HMI tags "New_Added"
   "AbufferCopyCut" : Bool, internal
   "AbufferFile" : WString[255], internal
   "AbufferFolder" : WString[255], internal
   "AbufferIsFolder" : Bool, internal
   "AFEsearchFolder" : WString[80], internal
   "AFEsearchString" : WString[80], internal
   "AFEStatus" : WString[150], internal
   "AFile_1" : WString[255], internal
   "AFile_10" : WString[255], internal
   "AFile_2" : WString[255], internal
   "AFile_3" : WString[255], internal
   "AFile_4" : WString[255], internal
   "AFile_5" : WString[255], internal
   "AFile_6" : WString[255], internal
   "AFile_7" : WString[255], internal
   "AFile_8" : WString[255], internal
   "AFile_9" : WString[255], internal
   "AfileChosen" : Int, internal
   "AFolder" : WString[255], internal
   "AhtmlPath" : WString[80], internal
   "Aindex" : Int, internal
   "AisFolder_1" : WString[10], internal
   "AisFolder_10" : WString[10], internal
   "AisFolder_2" : WString[10], internal
   "AisFolder_3" : WString[10], internal
   "AisFolder_4" : WString[10], internal
   "AisFolder_5" : WString[10], internal
   "AisFolder_6" : WString[10], internal
   "AisFolder_7" : WString[10], internal
   "AisFolder_8" : WString[10], internal
   "AisFolder_9" : WString[10], internal
   "ANewFolder" : WString[255], internal
   "ANewName" : WString[255], internal
   "ANextPossible" : Bool, internal
   "ApdfPath" : WString[80], internal
   "ASearch" : Bool, internal
   "AstateBackground" : Bool, internal
   "copyusb" : Bool, internal

HMI tags "NEW"
   "PV_1" : DInt AT %DB12.DBD32, 1 s
   "PV_2" : DInt AT %DB13.DBD28, 1 s
   "PV_3" : Int AT %DB12.DBW6, 1 s
   "SV_1" : DInt AT %DB16.DBD26, 1 s
   "SV_2" : Int AT %DB14.DBW20, 1 s
   "SV_3" : Int AT %DB12.DBW4, 1 s
   "Selection" : Bool AT %M30.0, 1 s
   "F2" : Bool AT %M30.1, 1 s
   "F3" : Bool AT %M33.3, 1 s
   "F4" : Bool AT %M33.4, 1 s
   "F5" : Bool AT %M30.3, 1 s
   "ON_OFF" : Bool AT %M30.1, 1 s
   "Indicator" : Bool AT %Q124.2, 1 s
   "F6" : Bool AT %M30.4, 1 s

discrete alarms
   1: 'All logs have been closed successfully.', class Sampling, trigger "Sampling_Alarm" bit 0
      on Coming: function_a9b64e44("Sampling_Alarm", 0)
   2: 'Log initialization ended. All logs OK.', class Sampling, trigger "Sampling_Alarm" bit 1
      on Coming: function_a9b64e44("Sampling_Alarm", 1)
   3: 'The log was successfully exported / The log was successfully exported to SD Card', class Sampling, trigger "Sampling_Alarm" bit 2
      on Coming: function_a9b64e44("Sampling_Alarm", 2)

text list "FLow_RPM": 0 'RPM'; 1 'FLOW RATE'

text list "ON_OFF": 0 'OFF'; 1 'ON'

graphic list "Nav_Recipe": 0 'labu1'; 1 'labu2'

graphic list "Check_Uncheck": 0 'images (7)'; 1 '_green_check.svg'

graphic list "pump": 2 'motor2'; 1 'motor'; 3 'motor'; 4 'motor2'; 5 'motor'; 6 'motor2'

graphic list "MH": 0 'graph'; 1 'graph - Copy'

graphic list "Home": 0 'images_3'; 1 'images - Copy'

graphic list "Scope": 0..12 'scope_1'; 13 'scope - Copy'; 14 'scope_1'

graphic list "oscilloscope": 0..8 'osiloskope'; 9 'osiloskope - Copy'; 10..14 'osiloskope'

graphic list "SelectorMenu": 0..10 's2_1'; 11 's2 - Copy'; 12..14 's2_1'

graphic list "Color": 0 'color1'; 1 'color1'; 2 'color3'; 4 'color5'; 8 'color6'; 16 'color7'

graphic list "SettingSys1": 0..6 'settingsys_1'; 7..13 'gear_setting'

graphic list "CleaningPiston": 0 'CleaningPistonX'; 1 'CleaningPiston'

graphic list "Tank_Sensor": 0 'PilotLight_Round_R_On_256c'; 1 'PilotLight_Round_G_On_256c'

graphic list "Circuit_Type": 0 'No mode'; 1 'Lowpress green'; 2 'lowpress circulation'; 3 'Reduced green'; 4 'Interval green'; 5 'high press circuit'; 6 'shot cycle'

graphic list "Operation Mode": 8 'No mode'; 1024 'manual mode'; 2048 'automatic mode'; 11 'barrel service'

graphic list "Print Function": 0 'printer off'; 1 'printer on'

graphic list "mh_switch_HP": 0 'blacklight'; 1 'greenlight'

graphic list "Nav_7": 0 'service solution'; 1..6 'gear_setting'

graphic list "icon_MHalarm": 1 'mixinghead_blue_alarm'; 2..15 'moxinghead_notblue_alarm'; 0 'moxinghead_notblue_alarm'

graphic list "icon_MHhyraulic": 0..1 'hydraulic_notblue_alarm'; 2 'hydraulic_blue_alarm'; 3..15 'hydraulic_notblue_alarm'

graphic list "ico_Pump": 0..2 'pump_notblue'; 3 'pump_blue'; 4..15 'pump_notblue'

graphic list "ico_machine": 0..4 'machine_notblue'; 5 'machine_blue'; 6..15 'machine_notblue'

graphic list "ico_alarm": 0 'alarmstate1'; 1 'alarmstate1_blue'; 2..20 'alarmstate1'

graphic list "ico_ShiftPlan": 0 'settingshiftplant1'; 1 'settingshiftplant2'; 2..5 'settingshiftplant1'

graphic list "ico_ShiftProtocol": 0..1 'ShiftProtocol1'; 2 'Shift_Protocol2'; 3..5 'ShiftProtocol1'

graphic list "ico_Actual_Fault": 0 'fault_2'; 1..3 'fault_1'

graphic list "ico_Actual_Fault_2": 0..10 'fault_1'; 11 'fault_2'; 12..15 'fault_1'

graphic list "ico_LastShot": 0..2 'lastshot_1'; 3 'lastshot_2'; 4..5 'lastshot_1'

graphic list "ico_Foaming": 0..1 'foaming_1'; 2 'foaming_2'; 3 'foaming_1'

graphic list "ico_Foaming_2": 0..11 'foaming_1'; 12 'foaming_2'; 13 'foaming_1'

graphic list "ico_ActualFault_Foaming": 0 'archiveFoam_1'; 1 'archiveFoam_2'; 2..15 'archiveFoam_1'

graphic list "ico_ActualFault_Foaming_2": 0..9 'archiveFoam_1'; 10 'archiveFoam_2'; 11..15 'archiveFoam_1'

graphic list "ico_MH": 0 'mixinghead_blue'; 1..2 'mixinghead_notblue'

graphic list "ico_Pump_large": 0 'pump_notblue'; 1 'pump_blue'; 2 'pump_notblue'

graphic list "ico_plcio": 9021 'plcio_2'; 9022..9024 'plcio1'; 9020 'plcio1'

graphic list "ico_consum": 0..3 'consumtion_1'; 4 'consumtion_2'; 5 'consumtion_1'

graphic list "Ico_navigation_2": 2 'Mcn_2'; 4 'mixinghead_blue'; 9 's2 - Copy'; 10 'Graphic_1'; 18 'process'; 21 'machine_2'; 24 'alarm_2'; 30 '021-online-learning-1'; 36 'lastshot_2'; 100 'scope - Copy'; 112 'Shift_Protocol2'; 113 'settingshiftplant2'; 887 'part counter_2'; 890 'consumtion_2'; 892 'chemical'; 999 '049-book'; 9020 'servicessolution_2'; 9021 'plcio_2'; 9024 'Graphic_29'; 15 'osiloskope - Copy'

graphic list "ico_information": 9020..9027 'information'; 9029 'information_2'

graphic list "@DiagnosticsStates": 0 '@Diagnostics_StateGood'; 1 '@Diagnostics_StateBad'

screen "0022_First_Screen" 1280x800, template "Navigation"
   TextField "KraussMaffei_Logo" at 289,360 size 714x81; Text 'Busur Kencana Sakti'
   TextField "KraussMaffei_Logo_1" at 434,435 size 328x47; Text 'POLYURETHANE'
   Button "first_btn" at 95,86 size 1084x711; TextOff '0017_Home Screen_OK'
      on Click: ActivateScreen("0017_Home Screen_OK", 0)

screen "0501_Trend_Sampling" 1280x800, template "Navigation"
   TextField "Text field_1" at 508,107 size 274x34; Text 'Trend Sampling Log'
   Button "print_2" at 1075,100 size 79x48; TextOff 'Text'; PictureOff "Graphic_10"
      on Click: function_f98d16b7()
      on Press: function_b14e0dd5("PrintScreenButton", 0)
      Appearance <- "PrintScreenButton"
   Rectangle "Rectangle_7" at 212,753 size 19x19
      Appearance <- "enable_poly_1"
   TextField "Text field_2" at 180,733 size 75x18; Text 'flowrate'
   Rectangle "Rectangle_9" at 284,753 size 19x19
      Appearance <- "enable_poly_2"
   TextField "Text field_13" at 257,733 size 73x18; Text 'pressure'
   Rectangle "Rectangle_1" at 348,753 size 19x19
      Appearance <- "enable_poly_3"
   TextField "Text field_4" at 332,733 size 63x18; Text 'Temp(C)'
   Rectangle "Rectangle_6" at 417,753 size 19x19
      Appearance <- "enable_poly_4"
   TextField "Text field_6" at 397,733 size 87x18; Text 'Speed (Rpm)'
   TextField "Text field_3" at 104,754 size 73x18; Text 'Poly'
   TextField "Text field_7" at 104,733 size 73x18; Text 'Ket.'
   FunctionTrendControl "f(x) trend view_1" at 103,151 size 1070x576
   Button "btn_safely" at 16,548 size 66x64; TextOn 'Safely'; TextOff 'Safely'; PictureOff "Graphic_16"; PictureList "ico_navigation_1"
      on Click: function_c6243368("safely_remove_usb", '\Storage Card USB\')
      ProcessValue <- "DB14_TP_Shortcuts_TP_Shortcuts_PageNo_7"

screen "0502_Trend Historical" 1280x800, template "Navigation"
   on GenerateScreen: SetTag("current_dir", '\Storage Card SD\Sampling\')
   TextField "Text field_1" at 471,107 size 348x34; Text 'Historical sampling trend'
   Button "pilih_file" at 986,744 size 77x38; TextOff '.... / ......'
      on Click: function_f12b67b1('*.csv*', '\Storage Card SD\Archive', 1, 1, 1, 1, "fileChossen", "stat_fileChosen")
   IOField "I/O field_1" at 489,746 size 478x39; FormatPattern ????????????????????????????????????????????????????????????????????????????????
      ProcessValue <- "fileChossen"
   Button "refresh_1" at 16,678 size 68x66; TextOff 'Refresh'; PictureOff "Graphic_22"
      on Click: function_bb0abc73(); ActivateScreen("0502_Trend Historical", 0)
   Button "open_file" at 1068,744 size 96x38; TextOff 'Open'
      on Click: function_efd5fb8c(); "Restore_Archive"()
      Appearance <- "Anim_OpenLOgs"
      on Press: function_b14e0dd5("Anim_OpenLOgs", 0)
   FunctionTrendControl "Trend_Log_view" at 103,151 size 1070x576
      TrendBeginTime <- "Trend_startingTime"
      TrendEndTime <- "Trend_endTime"
   Button "print_1" at 1075,100 size 79x48; TextOff 'Text'; PictureOff "Graphic_10"
      on Click: function_f98d16b7()
      on Press: function_b14e0dd5("PrintScreenButton", 0)
      Appearance <- "PrintScreenButton"
   Rectangle "Rectangle_7" at 212,753 size 19x19
      Appearance <- "enable_poly_1"
   TextField "Text field_2" at 180,733 size 75x18; Text 'flowrate'
   Rectangle "Rectangle_9" at 284,753 size 19x19
      Appearance <- "enable_poly_2"
   TextField "Text field_13" at 257,733 size 73x18; Text 'pressure'
   Rectangle "Rectangle_1" at 348,753 size 19x19
      Appearance <- "enable_poly_3"
   TextField "Text field_4" at 332,733 size 63x18; Text 'Temp(C)'
   Rectangle "Rectangle_6" at 417,753 size 19x19
      Appearance <- "enable_poly_4"
   TextField "Text field_6" at 397,733 size 87x18; Text 'Speed (Rpm)'
   TextField "Text field_3" at 104,754 size 73x18; Text 'Poly'
   TextField "Text field_7" at 104,733 size 73x18; Text 'Ket.'

screen "0500_Sampling Menu" 1280x800, template "Navigation"
   Button "save_data" at 113,167 size 203x60; TextOff 'SAVE DATA'
      on Click: InvertBit("saveDataControl")
      Appearance <- "saveDataControl"
   Button "log_data" at 370,167 size 203x60; TextOff 'LOG DATA'
      on Click: function_fd9437ed(0, "Current_Log"); InvertBit("loggingDataControl")
      Appearance <- "loggingDataControl"
   Button "clrrr" at 628,166 size 203x60; TextOff 'Clear'
      on Click: InvertBit("cleardata"); function_ff1151d2(0, "Current_Log"); SetTag("count", 0)
      Appearance <- "cleardata"
   Button "Closealllogs" at 113,265 size 203x60; TextOff 'Close All Logs'
      on Click: function_efd5fb8c()
   Button "openalllogs" at 370,265 size 203x60; TextOff 'Open All Logs'
      on Click: function_bb0abc73()
   Button "archive_log" at 628,265 size 203x60; TextOff 'Archive Log'
      on Click: function_e9be9208(0, "Current_Log", '\Storage Card SD\Archive', 0)
   Button "Button_12" at 113,364 size 203x60; TextOff 'File Explorer'
      on Click: SetTag("Folder", '\Storage Card SD\pdffile\'); SetTag("AFolder", '\Storage Card USB\'); ActivateScreen("0503_File_Explrr", 0)
   AlarmView "Alarm view_1" at 565,462 size 601x331
   TextField "Text field_2" at 497,107 size 295x34; Text 'Sampling Log Control'
   IOField "I/O field_1" at 937,221 size 146x59; FormatPattern 999
      ProcessValue <- "count"
   IOField "I/O field_2" at 935,334 size 146x56; FormatPattern 9999
      ProcessValue <- "Sampling_Time"
   TextField "Text field_1" at 937,186 size 173x25; Text 'Logging proggres'
   TextField "Text field_3" at 937,298 size 144x25; Text 'Sampling Time'
   TextField "Text field_4" at 1085,349 size 50x25; Text '[ms]'
   Button "sampling_trend" at 370,364 size 203x60; TextOff 'Sampling Trend'
      on Click: ActivateScreen("0501_Trend_Sampling", 0)
   Button "historical_sampl" at 628,364 size 203x60; TextOff 'Historical Sampling'
      on Click: ActivateScreen("0502_Trend Historical", 0)
   Button "clear_alrm" at 17,679 size 66x64; TextOff 'Text'; PictureOff "Graphic_14"
      on Click: function_e14cd482("Sampling")
   TextField "Text field_5" at 116,467 size 435x42; Text 'Enable Disable Logging data :'
   TextField "Text field_6" at 135,517 size 225x25; Text 'Flowrate'
   Button "check_enabletool" at 402,518 size 40x25; TextOff 'Text'; PictureList "Check_Uncheck"; PictureOff "download"
      on Click: InvertBit("enable_poly_1")
      ProcessValue <- "enable_poly_1"
   TextField "Text field_8" at 135,581 size 225x25; Text 'Pressure'
   Button "check_enabletool_2" at 402,582 size 40x25; TextOff 'Text'; PictureList "Check_Uncheck"; PictureOff "download"
      on Click: InvertBit("enable_poly_2")
      ProcessValue <- "enable_poly_2"
   TextField "Text field_10" at 135,645 size 225x25; Text 'Temperature'
   Button "check_enabletool_4" at 402,646 size 40x25; TextOff 'Text'; PictureList "Check_Uncheck"; PictureOff "download"
      on Click: InvertBit("enable_poly_3")
      ProcessValue <- "enable_poly_3"
   TextField "Text field_12" at 135,709 size 225x25; Text 'Rpm'
   Button "check_enabletool_6" at 402,710 size 40x25; TextOff 'Text'; PictureList "Check_Uncheck"; PictureOff "download"
      on Click: InvertBit("enable_poly_4")
      ProcessValue <- "enable_poly_4"
   Button "clear_alrm_1" at 1196,290 size 66x64; TextOff 'Text'; PictureOff "Graphic_32"
      on Click: ActivateScreen("Alarm", 0)

screen "LHmiView_FileExplorer" 1280x800, template "Navigation"
   on ClearScreen: ResetBit("stateBackground")
   on GenerateScreen: SetTag("Folder", '\Storage Card SD\')
   Button "btnDarkBackground" at 109,98 size 1062x681; TextOff 'Text'; PictureOff "Dark_Background"; PictureOn "Dark_Background"
      Visibility <- "stateBackground"
   TextField "Text field_2" at 130,107 size 177x34; Text 'File Explorer'
   Button "btnScrollUp" at 957,290 size 56x68; TextOff 'SPEICHERN / Open Path / SAVE'; PictureOff "Graphic_5"
      on Click: function_b9b71300("index", 1); "LHmiView_vbsFEWriteFilePropertiesToTags"("index")
      ObjectEnable <- "index"
   Button "btnScrollDown" at 957,630 size 56x68; TextOff 'SPEICHERN / Open Path / SAVE'; PictureOff "Graphic_6"
      on Click: function_dd21b452("index", 1); "LHmiView_vbsFEWriteFilePropertiesToTags"("index")
      ObjectEnable <- "NextPossible"
   Circle "Circle_1" at 972,170 size 29x29
      Appearance <- "copyusb"
   Button "de" at 951,159 size 66x49; TextOff 'Text'
      on Click: InvertBit("copyusb")
   TextField "txtFilter" at 137,251 size 56x24; Text 'Filter:'
   TextField "txtPath" at 137,199 size 56x24; Text 'Path: / Pfad:'
   Button "btn_safely" at 16,724 size 68x66; TextOn 'Safely'; TextOff 'Safely'; PictureOff "Graphic_16"; PictureList "ico_navigation_1"
      on Click: function_c6243368("safely_remove_usb", '\Storage Card USB\')
      ProcessValue <- "DB14_TP_Shortcuts_TP_Shortcuts_PageNo_7"
   Button "btn_safely_1" at 16,539 size 68x66; TextOn 'Safely'; TextOff 'Safely'; Authorization "Operate"; PictureOff "Graphic_21"; PictureList "ico_navigation_1"
      on Click: StopRuntime(0)
      ProcessValue <- "DB14_TP_Shortcuts_TP_Shortcuts_PageNo_7"
   IOField "ioPath" at 209,189 size 738x43; FormatPattern ??????????????????????????????????????????????????
      ProcessValue <- "Folder"
   IOField "ioFilter" at 209,241 size 738x43; FormatPattern ??????????????????????????????????????????????????
      ProcessValue <- "FEsearchString"
   Button "btnDeleteFilter" at 1061,170 size 72x50; TextOff 'Text'; PictureOff "Graphic_4"
      on Click: "LHmiView_vbsFEPreviousFolder"()
   Button "btnOpen" at 1061,228 size 72x50; TextOff 'Text'; PictureOn "Read"; PictureOff "Graphic_3"
      on Click: "LHmiView_vbsFEShowFiles"()
   Button "btnSearch" at 1061,287 size 72x50; TextOff 'Text'; PictureOn "Search"; PictureOff "Graphic_7"
      on Click: SetTag("Search", 1); "LHmiView_vbsFESearch"()
   Button "btnNew" at 1061,404 size 72x50; TextOff 'Text'; PictureOn "LHmiView_NewFolderFE"; PictureOff "LHmiView_NewFolderFE"
      on Click: function_efd93a16("LHmiView_popupFENewFolder", 432, 306, -1, -1, 1)
   Button "btnDelete" at 1061,345 size 72x50; TextOff 'Text'; PictureOn "LHmiView_DeleteFE"; PictureOff "LHmiView_DeleteFE"
      on Click: function_efd93a16("LHmiView_popupFEDelete", 432, 306, -1, -1, 1)
   Button "btnRename" at 1061,462 size 72x50; TextOff 'Text'; PictureOn "LHmiView_RenameFE"; PictureOff "LHmiView_RenameFE"
      on Click: function_efd93a16("LHmiView_popupFERename", 432, 306, -1, -1, 1)
   Button "btnCopy" at 1061,521 size 72x50; TextOff 'Text'; PictureOn "LHmiView_CopyFE"; PictureOff "LHmiView_CopyFE"
      on Click: "LHmiView_vbsFEMove"(1)
   Button "btnCut" at 1061,638 size 72x50; TextOff 'Text'; PictureOn "Link_White_26_22"; PictureOff "Graphic_2"
      on Click: "LHmiView_vbsFEMove"(3)
   Button "btnPaste" at 1061,579 size 72x50; TextOff 'Text'; PictureOn "LHmiView_PasteFE"; PictureOff "LHmiView_PasteFE"
      on Click: "LHmiView_vbsFEMove"(2)
   IOField "ioFile10" at 143,653 size 808x43; FormatPattern ????????????????????????????????????????????????????????????????????????????????
      ProcessValue <- "File_10"
      Appearance <- "fileChosen"
   IOField "ioFile1" at 143,293 size 808x43; FormatPattern ????????????????????????????????????????????????????????????????????????????????
      ProcessValue <- "File_1"
      Appearance <- "fileChosen"
   IOField "ioFile2" at 143,333 size 808x43; FormatPattern ????????????????????????????????????????????????????????????????????????????????
      ProcessValue <- "File_2"
      Appearance <- "fileChosen"
   IOField "ioFile3" at 143,373 size 808x43; FormatPattern ????????????????????????????????????????????????????????????????????????????????
      ProcessValue <- "File_3"
      Appearance <- "fileChosen"
   IOField "ioFile4" at 143,413 size 808x43; FormatPattern ????????????????????????????????????????????????????????????????????????????????
      ProcessValue <- "File_4"
      Appearance <- "fileChosen"
   IOField "ioFile5" at 143,453 size 808x43; FormatPattern ????????????????????????????????????????????????????????????????????????????????
      ProcessValue <- "File_5"
      Appearance <- "fileChosen"
   IOField "ioFile6" at 143,493 size 808x43; FormatPattern ????????????????????????????????????????????????????????????????????????????????
      ProcessValue <- "File_6"
      Appearance <- "fileChosen"
   IOField "ioFile7" at 143,533 size 808x43; FormatPattern ????????????????????????????????????????????????????????????????????????????????
      ProcessValue <- "File_7"
      Appearance <- "fileChosen"
   IOField "ioFile8" at 143,573 size 808x43; FormatPattern ????????????????????????????????????????????????????????????????????????????????
      ProcessValue <- "File_8"
      Appearance <- "fileChosen"
   IOField "ioFile9" at 143,613 size 808x43; FormatPattern ????????????????????????????????????????????????????????????????????????????????
      ProcessValue <- "File_9"
      Appearance <- "fileChosen"
   Button "btnFile1" at 142,293 size 809x43; TextOff 'Text'
      on Click: SetTag("fileChosen", 1)
   Button "btnFile2" at 142,333 size 809x43; TextOff 'Text'
      on Click: SetTag("fileChosen", 2)
   Button "btnFile3" at 142,373 size 809x43; TextOff 'Text'
      on Click: SetTag("fileChosen", 3)
   Button "btnFile4" at 142,413 size 809x43; TextOff 'Text'
      on Click: SetTag("fileChosen", 4)
   Button "btnFile5" at 142,453 size 809x43; TextOff 'Text'
      on Click: SetTag("fileChosen", 5)
   Button "btnFile6" at 142,493 size 809x43; TextOff 'Text'
      on Click: SetTag("fileChosen", 6)
   Button "btnFile7" at 142,533 size 809x43; TextOff 'Text'
      on Click: SetTag("fileChosen", 7)
   Button "btnFile8" at 142,573 size 809x43; TextOff 'Text'
      on Click: SetTag("fileChosen", 8)
   Button "btnFile9" at 142,613 size 809x43; TextOff 'Text'
      on Click: SetTag("fileChosen", 9)
   Button "btnFile10" at 142,653 size 809x43; TextOff 'Text'
      on Click: SetTag("fileChosen", 10)
   TextField "txtSate" at 183,733 size 913x24; Text 'State: / Status: / Status :'

screen "0503_File_Explrr" 1280x800, template "Navigation"
   on ClearScreen: ResetBit("AstateBackground"); ResetBit("stateBackground")
   on GenerateScreen: SetBit("copyusb")
   TextField "Text field_2" at 130,107 size 226x34; Text 'Managemen File'
   Button "btnScrollUp" at 580,253 size 56x68; TextOff 'SPEICHERN / Open Path / SAVE'; PictureOff "Graphic_5"
      on Click: function_b9b71300("index", 1); "LHmiView_vbsFEWriteFilePropertiesToTags"("index")
      ObjectEnable <- "index"
   Button "btnScrollDown" at 580,593 size 56x68; TextOff 'SPEICHERN / Open Path / SAVE'; PictureOff "Graphic_6"
      on Click: function_dd21b452("index", 1); "LHmiView_vbsFEWriteFilePropertiesToTags"("index")
      ObjectEnable <- "NextPossible"
   Button "btnScrollUp_1" at 1116,253 size 56x68; TextOff 'SPEICHERN / Open Path / SAVE'; PictureOff "Graphic_5"
      on Click: function_b9b71300("Aindex", 1); "LHmiView_vbsFEWriteFilePropertiesToTags_1"("Aindex")
      ObjectEnable <- "Aindex"
   Button "btnScrollDown_1" at 1116,593 size 56x68; TextOff 'SPEICHERN / Open Path / SAVE'; PictureOff "Graphic_6"
      on Click: function_dd21b452("Aindex", 1); "LHmiView_vbsFEWriteFilePropertiesToTags_1"("Aindex")
      ObjectEnable <- "ANextPossible"
   Button "file_explrr" at 16,290 size 65x63; TextOn 'Screen_2'; TextOff 'Screen_2'
      on Click: ActivateScreen("LHmiView_FileExplorer", 0)
   Button "explrer" at 1041,105 size 128x41; TextOff 'explorer.exe'
      on Click: function_bf5b406f('explorer.exe', '', 0, 0)
   IOField "ioPath" at 172,167 size 391x43; FormatPattern ??????????????????????????????????????????????????
      ProcessValue <- "Folder"
   IOField "ioFilter" at 172,219 size 391x43; FormatPattern ??????????????????????????????????????????????????
      ProcessValue <- "FEsearchString"
   IOField "ioPath_1" at 716,167 size 393x43; FormatPattern ??????????????????????????????????????????????????
      ProcessValue <- "AFolder"
   IOField "ioFilter_1" at 716,219 size 393x43; FormatPattern ??????????????????????????????????????????????????
      ProcessValue <- "AFEsearchString"
   TextField "txtFilter" at 105,229 size 49x25; Text 'Filter:'
   TextField "txtPath" at 105,177 size 44x25; Text 'Path: / Pfad:'
   TextField "txtFilter_1" at 649,229 size 49x25; Text 'Filter:'
   TextField "txtPath_1" at 649,177 size 44x25; Text 'Path: / Pfad:'
   Button "btn_safely" at 16,678 size 68x66; TextOn 'Safely'; TextOff 'Safely'; PictureOff "Graphic_16"; PictureList "ico_navigation_1"
      on Click: function_c6243368("safely_remove_usb", '\Storage Card USB\')
      ProcessValue <- "DB14_TP_Shortcuts_TP_Shortcuts_PageNo_7"
   Button "btn_safely_1" at 16,548 size 68x66; TextOn 'Safely'; TextOff 'Safely'; PictureOff "Graphic_21"; PictureList "ico_navigation_1"
      on Click: StopRuntime(0)
      ProcessValue <- "DB14_TP_Shortcuts_TP_Shortcuts_PageNo_7"
   IOField "ioFile10" at 106,631 size 468x43; FormatPattern ????????????????????????????????????????????????????????????????????????????????
      ProcessValue <- "File_10"
      Appearance <- "fileChosen"
   IOField "ioFile1" at 106,271 size 468x43; FormatPattern ????????????????????????????????????????????????????????????????????????????????
      ProcessValue <- "File_1"
      Appearance <- "fileChosen"
   IOField "ioFile2" at 106,311 size 468x43; FormatPattern ????????????????????????????????????????????????????????????????????????????????
      ProcessValue <- "File_2"
      Appearance <- "fileChosen"
   IOField "ioFile3" at 106,351 size 468x43; FormatPattern ????????????????????????????????????????????????????????????????????????????????
      ProcessValue <- "File_3"
      Appearance <- "fileChosen"
   IOField "ioFile4" at 106,391 size 468x43; FormatPattern ????????????????????????????????????????????????????????????????????????????????
      ProcessValue <- "File_4"
      Appearance <- "fileChosen"
   IOField "ioFile5" at 106,431 size 468x43; FormatPattern ????????????????????????????????????????????????????????????????????????????????
      ProcessValue <- "File_5"
      Appearance <- "fileChosen"
   IOField "ioFile6" at 106,471 size 468x43; FormatPattern ????????????????????????????????????????????????????????????????????????????????
      ProcessValue <- "File_6"
      Appearance <- "fileChosen"
   IOField "ioFile7" at 106,511 size 468x43; FormatPattern ????????????????????????????????????????????????????????????????????????????????
      ProcessValue <- "File_7"
      Appearance <- "fileChosen"
   IOField "ioFile8" at 106,551 size 468x43; FormatPattern ????????????????????????????????????????????????????????????????????????????????
      ProcessValue <- "File_8"
      Appearance <- "fileChosen"
   IOField "ioFile9" at 106,591 size 468x43; FormatPattern ????????????????????????????????????????????????????????????????????????????????
      ProcessValue <- "File_9"
      Appearance <- "fileChosen"
   IOField "ioFile10_1" at 642,631 size 469x43; FormatPattern ????????????????????????????????????????????????????????????????????????????????
      ProcessValue <- "AFile_10"
      Appearance <- "AfileChosen"
   IOField "ioFile1_1" at 642,271 size 469x43; FormatPattern ????????????????????????????????????????????????????????????????????????????????
      ProcessValue <- "AFile_1"
      Appearance <- "AfileChosen"
   IOField "ioFile2_1" at 642,311 size 469x43; FormatPattern ????????????????????????????????????????????????????????????????????????????????
      ProcessValue <- "AFile_2"
      Appearance <- "AfileChosen"
   IOField "ioFile3_1" at 642,351 size 469x43; FormatPattern ????????????????????????????????????????????????????????????????????????????????
      ProcessValue <- "AFile_3"
      Appearance <- "AfileChosen"
   IOField "ioFile4_1" at 642,391 size 469x43; FormatPattern ????????????????????????????????????????????????????????????????????????????????
      ProcessValue <- "AFile_4"
      Appearance <- "AfileChosen"
   IOField "ioFile5_1" at 642,431 size 469x43; FormatPattern ????????????????????????????????????????????????????????????????????????????????
      ProcessValue <- "AFile_5"
      Appearance <- "AfileChosen"
   IOField "ioFile6_1" at 642,471 size 469x43; FormatPattern ????????????????????????????????????????????????????????????????????????????????
      ProcessValue <- "AFile_6"
      Appearance <- "AfileChosen"
   IOField "ioFile7_1" at 642,511 size 469x43; FormatPattern ????????????????????????????????????????????????????????????????????????????????
      ProcessValue <- "AFile_7"
      Appearance <- "AfileChosen"
   IOField "ioFile8_1" at 642,551 size 469x43; FormatPattern ????????????????????????????????????????????????????????????????????????????????
      ProcessValue <- "AFile_8"
      Appearance <- "AfileChosen"
   IOField "ioFile9_1" at 642,591 size 469x43; FormatPattern ????????????????????????????????????????????????????????????????????????????????
      ProcessValue <- "AFile_9"
      Appearance <- "AfileChosen"
   Button "btnFile1" at 105,271 size 468x43; TextOff 'Text'
      on Click: SetTag("fileChosen", 1)
   Button "btnFile2" at 105,311 size 468x43; TextOff 'Text'
      on Click: SetTag("fileChosen", 2)
   Button "btnFile3" at 105,351 size 468x43; TextOff 'Text'
      on Click: SetTag("fileChosen", 3)
   Button "btnFile4" at 105,391 size 468x43; TextOff 'Text'
      on Click: SetTag("fileChosen", 4)
   Button "btnFile5" at 105,431 size 468x43; TextOff 'Text'
      on Click: SetTag("fileChosen", 5)
   Button "btnFile6" at 105,471 size 468x43; TextOff 'Text'
      on Click: SetTag("fileChosen", 6)
   Button "btnFile7" at 105,511 size 468x43; TextOff 'Text'
      on Click: SetTag("fileChosen", 7)
   Button "btnFile8" at 105,551 size 468x43; TextOff 'Text'
      on Click: SetTag("fileChosen", 8)
   Button "btnFile9" at 105,591 size 468x43; TextOff 'Text'
      on Click: SetTag("fileChosen", 9)
   Button "btnFile10" at 105,631 size 468x43; TextOff 'Text'
      on Click: SetTag("fileChosen", 10)
   Button "btnFile1_1" at 644,271 size 466x43; TextOff 'Text'
      on Click: SetTag("AfileChosen", 1)
   Button "btnFile2_1" at 644,311 size 466x43; TextOff 'Text'
      on Click: SetTag("AfileChosen", 2)
   Button "btnFile3_1" at 644,351 size 466x43; TextOff 'Text'
      on Click: SetTag("AfileChosen", 3)
   Button "btnFile4_1" at 644,391 size 466x43; TextOff 'Text'
      on Click: SetTag("AfileChosen", 4)
   Button "btnFile5_1" at 644,431 size 466x43; TextOff 'Text'
      on Click: SetTag("AfileChosen", 5)
   Button "btnFile6_1" at 644,471 size 466x43; TextOff 'Text'
      on Click: SetTag("AfileChosen", 6)
   Button "btnFile7_1" at 644,511 size 466x43; TextOff 'Text'
      on Click: SetTag("AfileChosen", 7)
   Button "btnFile8_1" at 644,551 size 466x43; TextOff 'Text'
      on Click: SetTag("AfileChosen", 8)
   Button "btnFile9_1" at 644,591 size 466x43; TextOff 'Text'
      on Click: SetTag("AfileChosen", 9)
   Button "btnFile10_1" at 644,631 size 466x43; TextOff 'Text'
      on Click: SetTag("AfileChosen", 10)
   TextField "txtSate" at 117,740 size 1031x24; Text 'State: / Status: / Message :'
   TextField "txtSate_1" at 117,765 size 1032x24; Text 'State: / Status: / Message :'
   Rectangle "Rectangle_4" at 104,675 size 481x59
      Visibility <- "CopyfromUSB"
   Rectangle "Rectangle_3" at 640,676 size 481x59
      Visibility <- "CopyfromSD"
   Button "btnDeleteFilter" at 107,680 size 72x50; TextOff 'Text'; PictureOff "Graphic_4"
      on Click: "LHmiView_vbsFEPreviousFolder"()
   Button "btnOpen" at 185,680 size 72x50; TextOff 'Text'; PictureOn "Read"; PictureOff "Graphic_3"
      on Click: "LHmiView_vbsFEShowFiles"()
   Button "btnSearch" at 263,680 size 72x50; TextOff 'Text'; PictureOn "Search"; PictureOff "Graphic_7"
      on Click: SetTag("Search", 1); "LHmiView_vbsFESearch"()
   Button "btnDeleteFilter_1" at 644,680 size 72x50; TextOff 'Text'; PictureOff "Graphic_4"
      on Click: "LHmiView_vbsFEPreviousFolder_1"()
   Button "btnOpen_1" at 722,680 size 72x50; TextOff 'Text'; PictureOn "Read"; PictureOff "Graphic_3"
      on Click: "LHmiView_vbsFEShowFiles_1"()
   Button "btnSearch_1" at 801,680 size 72x50; TextOff 'Text'; PictureOn "Search"; PictureOff "Graphic_7"
      on Click: SetTag("ASearch", 1); "LHmiView_vbsFESearch_1"()
   Button "btnCopy" at 419,680 size 72x50; TextOff 'Text'; PictureOn "LHmiView_CopyFE"; PictureOff "LHmiView_CopyFE"
      on Click: "LHmiView_vbsFEMove_1"(1); SetBit("CopyfromSD")
      Visibility <- "copyusb"
   Button "btnPaste" at 498,680 size 72x50; TextOff 'Text'; PictureOn "LHmiView_PasteFE"; PictureOff "LHmiView_PasteFE"
      on Click: "LHmiView_vbsFEMove_1"(2); ResetBit("CopyfromSD")
      Visibility <- "copyusb"
   Button "btnDelete" at 341,680 size 72x50; TextOff 'Text'; PictureOn "LHmiView_DeleteFE"; PictureOff "LHmiView_DeleteFE"
      on Click: function_efd93a16("LHmiView_popupFEDelete_2", 189, 332, -1, -1, 1)
   Button "btnDelete_1" at 879,680 size 72x50; TextOff 'Text'; PictureOn "LHmiView_DeleteFE"; PictureOff "LHmiView_DeleteFE"
      on Click: function_efd93a16("LHmiView_popupFEDelete_1", 713, 332, -1, -1, 1)
   Button "btnCopy_1" at 958,680 size 72x50; TextOff 'Text'; PictureOn "LHmiView_CopyFE"; PictureOff "LHmiView_CopyFE"
      on Click: "LHmiView_vbsFEMove"(1); SetBit("CopyfromUSB")
      Visibility <- "copyusb"
   Button "btnPaste_1" at 1037,680 size 72x50; TextOff 'Text'; PictureOn "LHmiView_PasteFE"; PictureOff "LHmiView_PasteFE"
      on Click: "LHmiView_vbsFEMove"(2); ResetBit("CopyfromUSB")
      Visibility <- "copyusb"
   Button "btnPaste_2" at 572,164 size 72x50; TextOff 'Text'; PictureOn "LHmiView_PasteFE"; PictureOff "Graphic_20"
      on Click: "LHmiView_vbsFEReadFilesOfFolder"("Folder"); "LHmiView_vbsFEWriteFilePropertiesToTags"("index"); "LHmiView_vbsFEReadFilesOfFolder_1"("AFolder"); "LHmiView_vbsFEWriteFilePropertiesToTags_1"("Aindex")
   Button "btnCopy_2" at 419,680 size 72x50; TextOff 'Text'; PictureOn "LHmiView_CopyFE"; PictureOff "LHmiView_CopyFE"
      on Click: "LHmiView_vbsFEMove"(1); SetBit("CopyfromSD")
      Visibility <- "copyusb"
   Button "btnPaste_3" at 498,680 size 72x50; TextOff 'Text'; PictureOn "LHmiView_PasteFE"; PictureOff "LHmiView_PasteFE"
      on Click: "LHmiView_vbsFEMove"(2); ResetBit("CopyfromSD")
      Visibility <- "copyusb"
   Button "btnCopy_3" at 958,680 size 72x50; TextOff 'Text'; PictureOn "LHmiView_CopyFE"; PictureOff "LHmiView_CopyFE"
      on Click: "LHmiView_vbsFEMove_1"(1); SetBit("CopyfromUSB")
      Visibility <- "copyusb"
   Button "btnPaste_4" at 1037,680 size 72x50; TextOff 'Text'; PictureOn "LHmiView_PasteFE"; PictureOff "LHmiView_PasteFE"
      on Click: "LHmiView_vbsFEMove_1"(2); ResetBit("CopyfromUSB")
      Visibility <- "copyusb"
   Button "btnDarkBackground" at 1,4 size 650x795; TextOff 'Text'; PictureOn "Dark_Background"; PictureOff "Dark_Background"
      Visibility <- "stateBackground"
   Button "btnDarkBackground_1" at 630,4 size 650x795; TextOff 'Text'; PictureOff "Dark_Background"; PictureOn "Dark_Background"
      Visibility <- "AstateBackground"

Template "Navigation" 1280x800
   TextField "Template_Text field_1" at 1043,13 size 216x64; Text 'Busur Kencana Sakti'
   DateTimeField "Template_Date/time field_1" at 103,25 size 273x28
   Button "Button_7" at 16,15 size 66x48; TextOff 'BACK'; PictureOff "Graphic_4"
      on Click: function_efd93a16()
   Button "Button_6" at 16,678 size 66x64; TextOff 'Text'; PictureOff "Graphic_26"
      on Click: ActivateScreen("iNFO", 0)
   Button "Button_1" at 16,548 size 66x64; TextOff 'Text'; PictureOff "Graphic_14"
   Button "Button_2" at 16,419 size 66x64; TextOff 'Text'; PictureOff "Graphic_25"
      on Click: SetTag("Folder", '\Storage Card SD\pdffile\'); SetTag("AFolder", '\Storage Card USB\'); ActivateScreen("0503_File_Explrr", 0)
   Button "Button_3" at 16,290 size 66x64; TextOff 'Text'; PictureOff "Graphic_14"
   Button "Button_4" at 16,161 size 66x64; TextOff 'Text'; PictureOff "Graphic_24"
      on Click: ActivateScreen("0500_Sampling Menu", 0)
   Button "Button_5" at 1196,678 size 66x64; TextOff 'Text'; PictureOff "Graphic_30"
      on Click: ActivateScreen("0017_Home Screen_OK", 0)
   Button "Button_8" at 1196,548 size 66x64; TextOff 'Text'; PictureOff "Graphic_9"
   Button "Button_9" at 1196,419 size 66x64; TextOff 'Text'; PictureOff "Graphic_27"
      on Click: ActivateScreen("0502_Trend Historical", 0)
   Button "Button_10" at 1196,290 size 66x64; TextOff 'Text'; PictureOff "Graphic_8"
   Button "Button_11" at 1196,161 size 66x64; TextOff 'Text'; PictureOff "Graphic_8"
      on Click: ActivateScreen("0501_Trend_Sampling", 0)
   TextField "Template_Text field_2" at 668,20 size 137x39; Text 'Text'
      Appearance <- "Selection"
   TextField "Template_Text field_3" at 812,20 size 79x39; Text 'Text'
      Appearance <- "ON_OFF"
   TextField "Template_Text field_5" at 555,20 size 106x39; Text 'LOG DATA'
      Appearance <- "loggingDataControl"
   TextField "Template_Text field_6" at 434,20 size 114x39; Text 'SAVE DATA'
      Appearance <- "saveDataControl"
   Group "Group" at 898,20 size 50x39
   TextField "Template_Text field_7" at 555,20 size 106x39; Text 'LOG DATA'
      Visibility <- "loggingDataControl"
   TextField "Template_Text field_8" at 434,20 size 114x39; Text 'SAVE DATA'
      Visibility <- "saveDataControl"
   TextField "Template_Text field_4" at 898,20 size 50x39; Text 'Text'
   Circle "Template_Circle_1" at 909,26 size 28x28
      Appearance <- "Indicator"

PopupScreen "Sampling Popup" 500x300
   TextField "Text field_1" at 0,0 size 500x35; Text 'Log Control'
   Button "Button_4" at 455,3 size 43x32; TextOff 'X'
      on Click: function_efd93a16("Sampling Popup", 0, 0, 0, -1, 1)
   Button "Button_8" at 32,49 size 203x42; TextOff 'SAVE DATA'
      on Click: InvertBit("saveDataControl")
      Appearance <- "saveDataControl"
   Button "Button_9" at 252,49 size 203x42; TextOff 'LOG DATA'
      on Click: InvertBit("loggingDataControl")
      Appearance <- "loggingDataControl"
   Button "Button_10" at 87,113 size 311x42; TextOff 'Clear'
      on Click: InvertBit("cleardata"); function_ff1151d2(0, "Current_Log"); SetTag("count", 0)
      Appearance <- "cleardata"
   Button "Button_2" at 32,175 size 203x42; TextOff 'Close All Logs'
      on Click: function_efd5fb8c()
   Button "Button_3" at 252,175 size 203x42; TextOff 'Open All Logs'
      on Click: function_bb0abc73()
   Button "Button_1" at 32,235 size 203x42; TextOff 'Archive Log'
      on Click: function_e9be9208(0, "Current_Log", '\Storage Card SD\Archive', 0)
   Button "Button_12" at 252,237 size 203x42; TextOff 'COPY to USB'
      on Click: function_e9be9208(0, "Current_Log", '\Storage Card USB\', 0)

PopupScreen "LHmiView_popupFEDelete" 320x266
   on ClearScreen: ResetBit("stateBackground")
   on GenerateScreen: SetBit("stateBackground")
   TextField "Template_Text field_1" at 16,0 size 288x40; Text 'Delete file / folder / Datei / Ordner löschen / Delete File / Folder'
   Button "Button_2" at 16,210 size 288x40; TextOn 'CANCEL / ABBRECHEN'; TextOff 'CANCEL / ABBRECHEN'
      on Click: function_efd93a16("LHmiView_popupFEDelete", 0, 0, -1, -1, 1)
   Button "Schaltfläche_1" at 16,154 size 288x40; TextOn 'APPLY / BESTÄTIGEN'; TextOff 'BESTÄTIGEN / APPLY / YES'
      on Click: "LHmiView_vbsFEDelete"(); ActivateScreen("LHmiView_FileExplorer", 0)
   TextField "Text field_1" at 32,93 size 256x48; Text 'Do you really want to delete the file / folder? Wollen Sie die Datei / den Ordner wirklich löschen?'
   TextField "Text field_2" at 32,56 size 256x24; Text 'NOTE / HINWEIS / NOTE !!!'

PopupScreen "LHmiView_popupFENewFolder" 320x266
   on ClearScreen: ResetBit("stateBackground")
   on GenerateScreen: SetBit("stateBackground")
   TextField "txtChapter" at 16,0 size 288x40; Text 'Add new folder / Neuen Ordner hinzufügen'
   TextField "Text field_2" at 16,56 size 256x24; Text 'Name of new folder / Name neuer Ordner'
   IOField "ioNewFolder" at 16,82 size 288x40; FormatPattern ????????????????????????????????????????????????????????????????????????????????
      ProcessValue <- "NewFolder"
   Button "btnCancel" at 16,210 size 288x40; TextOff 'CANCEL / ABBRECHEN'
      on Click: ActivateScreen("LHmiView_FileExplorer", 0)
   Button "btnAdd" at 16,154 size 288x40; TextOn 'ADD / HINZUFÜGEN'; TextOff 'HINZUFÜGEN / ADD / YES'
      on Click: "LHmiView_vbsFECreateFolder"(); ActivateScreen("LHmiView_FileExplorer", 0)

PopupScreen "LHmiView_popupFERename" 320x266
   on ClearScreen: ResetBit("stateBackground")
   on GenerateScreen: SetBit("stateBackground")
   TextField "txtChapter" at 16,0 size 288x40; Text 'Rename file / folder / Datei / Ordner umbenennen'
   TextField "Text field_2" at 16,56 size 256x24; Text 'New name of file / folder / Neuer Name Datei / Ordner'
   IOField "ioNewFolder" at 16,82 size 288x40; FormatPattern ????????????????????????????????????????????????????????????????????????????????
      ProcessValue <- "NewName"
   Button "btnCancel" at 16,210 size 288x40; TextOff 'CANCEL / ABBRECHEN'
      on Click: ActivateScreen("LHmiView_FileExplorer", 0)
   Button "btnAdd" at 16,154 size 288x40; TextOn 'RENAME / UMBENNENEN'; TextOff 'UMBENNENEN / RENAME / YES'
      on Click: "LHmiView_vbsFERename"(); ActivateScreen("LHmiView_FileExplorer", 0)

PopupScreen "LHmiView_popupFEDelete_1" 320x266
   on ClearScreen: ResetBit("AstateBackground")
   on GenerateScreen: SetBit("AstateBackground")
   TextField "Template_Text field_1" at 16,0 size 288x40; Text 'Delete file / folder / Datei / Ordner löschen / Delete File / Folder'
   Button "Button_2" at 16,210 size 288x40; TextOn 'CANCEL / ABBRECHEN'; TextOff 'CANCEL / ABBRECHEN'
      on Click: function_efd93a16("LHmiView_popupFEDelete_1", 0, 0, -1, -1, 1)
   Button "Schaltfläche_1" at 16,154 size 288x40; TextOn 'APPLY / BESTÄTIGEN'; TextOff 'BESTÄTIGEN / APPLY / YES'
      on Click: "LHmiView_vbsFEDelete_1"(); ActivateScreen("0503_File_Explrr", 0)
   TextField "Text field_1" at 32,93 size 256x48; Text 'Do you really want to delete the file / folder? Wollen Sie die Datei / den Ordner wirklich löschen?'
   TextField "Text field_2" at 32,56 size 256x24; Text 'NOTE / HINWEIS / NOTE !!!'

PopupScreen "LHmiView_popupFEDelete_2" 320x266
   on ClearScreen: ResetBit("stateBackground")
   on GenerateScreen: SetBit("stateBackground")
   TextField "Template_Text field_1" at 16,0 size 288x40; Text 'Delete file / folder / Datei / Ordner löschen / Delete File / Folder'
   Button "Button_2" at 16,210 size 288x40; TextOn 'CANCEL / ABBRECHEN'; TextOff 'CANCEL / ABBRECHEN'
      on Click: function_efd93a16("LHmiView_popupFEDelete_2", 0, 0, -1, -1, 1)
   Button "Schaltfläche_1" at 16,154 size 288x40; TextOn 'APPLY / BESTÄTIGEN'; TextOff 'BESTÄTIGEN / APPLY / YES'
      on Click: "LHmiView_vbsFEDelete"(); ActivateScreen("0503_File_Explrr", 0)
   TextField "Text field_1" at 32,93 size 256x48; Text 'Do you really want to delete the file / folder? Wollen Sie die Datei / den Ordner wirklich löschen?'
   TextField "Text field_2" at 32,56 size 256x24; Text 'NOTE / HINWEIS / NOTE !!!'

screen "0017_Home Screen_OK" 1280x800, template "Navigation"
   on ClearScreen: SetTag("NavScreenChange", 0)
   IOField "I/O field_1" at 124,385 size 253x65; FormatPattern 99999
      ProcessValue <- "PV_1"
   IOField "I/O field_2" at 124,459 size 253x65; FormatPattern 99999
      ProcessValue <- "PV_2"
   IOField "I/O field_3" at 124,532 size 253x65; FormatPattern 99999
      ProcessValue <- "PV_3"
   IOField "I/O field_4" at 812,385 size 253x65; FormatPattern 99999
      ProcessValue <- "SV_1"
   IOField "I/O field_5" at 812,459 size 253x65; FormatPattern 99999
      ProcessValue <- "SV_2"
   IOField "I/O field_6" at 812,532 size 253x65; FormatPattern 99999
      ProcessValue <- "SV_3"
   TextField "Text field_2" at 813,283 size 342x70; Text 'SV'
   Button "pilihan" at 465,118 size 350x119; TextOff 'Text'; TextList "FLow_RPM"
      ProcessValue <- "Selection"
      on Click: InvertBit("Selection")
      Appearance <- "Selection"
   Button "n_f" at 526,340 size 228x85; TextOff 'Text'; TextList "ON_OFF"
      ProcessValue <- "ON_OFF"
      Appearance <- "ON_OFF"
      on Click: InvertBit("ON_OFF")
   Circle "Circle_1" at 586,488 size 108x108
      Appearance <- "Indicator"
   Button "up_2" at 465,661 size 132x95; TextOn 'UP'; TextOff 'UP'; TextList "ON_OFF"; PictureOff "Graphic_5"
      ProcessValue <- "ON_OFF"
      on Press: function_b14e0dd5("F5", 0)
      Appearance <- "F5"
      Visibility <- "Selection"
   Button "dwn_2" at 683,661 size 132x95; TextOff 'DOWN'; TextList "ON_OFF"; PictureOff "Graphic_6"
      on Press: function_b14e0dd5("F6", 0)
      ProcessValue <- "ON_OFF"
      Appearance <- "F6"
      Visibility <- "Selection"
   TextField "Text field_3" at 386,396 size 62x43; Text 'g/s'
   TextField "Text field_4" at 386,470 size 61x43; Text 'bar'
   TextField "Text field_5" at 386,543 size 45x43; Text '°C'
   TextField "Text field_6" at 1074,396 size 62x43; Text 'g/s'
   TextField "Text field_7" at 1074,470 size 73x43; Text 'rpm'
   TextField "Text field_8" at 1074,543 size 45x43; Text '°C'
   TextField "Text field_9" at 124,283 size 342x70; Text 'PV'
   Button "up_1" at 465,661 size 132x95; TextOn 'UP'; TextOff 'UP'; TextList "ON_OFF"; PictureOff "Graphic_5"
      on Press: function_b14e0dd5("F3", 0)
      ProcessValue <- "ON_OFF"
      Visibility <- "Selection"
      Appearance <- "F3"
   Button "dwn_1" at 683,661 size 132x95; TextOff 'DOWN'; PictureOff "Graphic_6"; TextList "ON_OFF"
      on Press: function_b14e0dd5("F4", 0)
      ProcessValue <- "ON_OFF"
      Visibility <- "Selection"
      Appearance <- "F4"

screen "iNFO" 1280x800, template "Navigation"
   Button "btn_safely_1" at 16,548 size 68x66; TextOn 'Safely'; TextOff 'Safely'; PictureOff "Graphic_21"; PictureList "ico_navigation_1"
      on Click: StopRuntime(0)
      ProcessValue <- "DB14_TP_Shortcuts_TP_Shortcuts_PageNo_7"
   TextField "Text field_1" at 367,197 size 203x40; Text 'Save Data'
   TextField "Text field_2" at 367,292 size 203x40; Text 'Log Data'
   TextField "Text field_3" at 367,387 size 203x40; Text 'Log Count = 600'
   TextField "Text field_4" at 367,482 size 203x40; Text 'Close All Logs'
   TextField "Text field_5" at 367,577 size 203x40; Text 'Archive Log'
   TextField "Text field_6" at 367,672 size 203x40; Text 'Open All Logs'
   TextField "Text field_7" at 163,130 size 230x40; Text 'Process Sampling Data'
   TextField "Text field_8" at 762,170 size 68x34; Text 'Date'
   DateTimeField "Date/time field_1" at 768,213 size 291x48
   DateTimeField "Date/time field_2" at 768,340 size 291x48
   TextField "Text field_9" at 762,299 size 71x34; Text 'Time'

screen "Alarm" 1280x800, template "Navigation"
   AlarmView "Alarm view_1" at 140,124 size 1000x640

VB script "StartStopLogging"
   If SmartTags("count") >= 600 Then
   	b6526003-1e6c-4105-b1c3-8571bad56740 $3$hmiDataLog$,Current_Log
   End If

VB script "Restore_Archive"
   'Tip:
   ' 1. Verwenden Sie die Tastenkombination <CTRL+SPACE> oder <CTRL+I>, um eine Liste aller Objekte und Funktionen zu öffnen
   ' 2. Schreiben Sie den Code unter Verwendung des HMI Runtime Objekts.
   '  Beispiel: HmiRuntime.Screens("Screen_1").
   ' 3. Verwenden Sie die Tastenkombination <CTRL+J>, um eine Objektreferenz zu erstellen.
   'Schreiben Sie den Code ab dieser Position:
   	Dim fs, f, f2
   	Dim source_name1, target_name1
   	Dim source_name2, target_name2
   	Dim source_name3, target_name3
   	Dim source_name4, target_name4
   	Dim source_name5, target_name5
   	Dim source_name6, target_name6
   	Dim source_name7, target_name7
   	Dim source_name8, target_name8
   	Dim source_name9, target_name9
   	Dim lta_path, lta_time, current_path				' "lta" = "long-term archive"
   	
   	' take the variable names, and enclose them in quotes:
   	source_name1= """" & "pressure_poly" & """"
   	target_name1= """" & "pressure_poly_res" & """"
   	source_name2= """" & "count" & """"
   	target_name2= """" & "count_res" & """"
   	source_name3= """" & "flowrate_poly" & """"
   	target_name3= """" & "flowrate_poly_res" & """"
   	source_name4= """" & "pressure_iso" & """"
   	target_name4= """" & "pressure_iso_res" & """"
   	source_name5= """" & "flowrate_iso" & """"
   	target_name5= """" & "flowrate_iso_res" & """"
   	source_name6= """" & "temperature_poly" & """"
   	target_name6= """" & "temperature_poly_res" & """"
   	source_name7= """" & "temperature_iso" & """"
   	target_name7= """" & "temperature_iso_res" & """"
   	source_name8= """" & "speed_poly" & """"
   	target_name8= """" & "speed_poly_res" & """"
   	source_name9= """" & "speed_iso" & """"
   	target_name9= """" & "speed_iso_res" & """"
   	
   	
   	Dim restore_entry, restore_fields
   	lta_path = SmartTags("fileChossen")
   	archive_path= lta_path
       current_path= current_dir & "RestoredLog0.csv"
       
   	Set fs = CreateObject("FileCtl.FileSystem") 	
   	bfde4b54-0db7-4817-8032-87127bf19bb9("Exploring <" & lta_path & ">, <" & current_path & ">.")
   	
   	' does the long-term archive exist?
   	If fs.Dir(lta_path)<>"" Then				' ***
   		
   		Set f= CreateObject("FileCtl.File")
   		Set f2= CreateObject("FileCtl.File")
   		
   	    f.Open current_path, 2			' write access, create if not existant
   		fs.setAttr lta_path, 0			' required on panels
   	    f2.Open lta_path, 1				' read access
   	
   		'---------------------------------------------------------
   		' the following code block is optional
   		' it extracts the date/time of the first archive data entry so the operator will have an idea
   		' when the archive was created:
   		' you can safely delete everything up to and including "End If"
   		
   	    restore_entry= f2.lineinputstring		' first line is no data point entry, copy to target:
   	    f.lineprint(restore_entry)
   	    restore_entry= f2.lineinputstring		' second line contains first data point, copy to target, too:
   			restore_entry= Replace(restore_entry, source_name1, target_name1)
   			restore_entry= Replace(restore_entry, source_name2, target_name2)
   			restore_entry= Replace(restore_entry, source_name3, target_name3)
   			restore_entry= Replace(restore_entry, source_name4, target_name4)
   			restore_entry= Replace(restore_entry, source_name5, target_name5)
   			restore_entry= Replace(restore_entry, source_name6, target_name6)
   			restore_entry= Replace(restore_entry, source_name7, target_name7)
   			restore_entry= Replace(restore_entry, source_name8, target_name8)
   			restore_entry= Replace(restore_entry, source_name9, target_name9)
   	    f.lineprint(restore_entry)
   	    
   	    ' extract date/time from this line (second entry in a CSV file):
   	    restore_fields= Split(restore_entry, ";")
   	    lta_time= Mid(restore_fields(1), 2, Len(restore_fields(1))-2)
   	    restore_time= CDate(Mid(restore_fields(1), 2, Len(restore_fields(1))-2))